VERSION : 0.1
   VAR_INPUT
      "array" : Variant;
   END_VAR
   VAR_TEMP
      status : DInt;
      ret : UDInt;
   END_VAR
BEGIN
   #ret := CountOfElements(#array);
   #"Array.Any.Length" := #ret;
END_FUNCTION

FUNCTION "Get Station Index From Id" : Int   // FC106, SCL
{ S7_Optimized_Access := 'TRUE' }
VERSION : 0.1
   VAR_INPUT
      line_name : WString;
      drop_zone : USInt;
      stns : "Station: All Stations";
   END_VAR
   VAR_TEMP
      i : Int;
      ret : Int;
   END_VAR
BEGIN
   REGION "MATCH LINE NAME AND DROP ZONE"
       FOR #i := 0 TO "STATION_COUNT" DO
           IF #line_name = #stns.stn[#i].id.lineName THEN
               IF #drop_zone = #stns.stn[#i].id.dropZone THEN
                   #ret := #i;
                   EXIT;
               END_IF;
           END_IF;
       END_FOR;
   END_REGION


   REGION "RETURN"
       #"Get Station Index From Id" := #ret;
   END_REGION
END_FUNCTION

FUNCTION "Array.Int.Fill" : Void   // FC109, SCL
{ S7_Optimized_Access := 'TRUE' }
VERSION : 0.1
   VAR_INPUT
      value : Int;
   END_VAR
   VAR_IN_OUT
      int_array : Array[*] of Int;
   END_VAR
   VAR_TEMP
      _i : DInt;
      _length : DInt;
   END_VAR
BEGIN
   REGION "GET LENGHT"
       #_length := UDINT_TO_DINT("Array.Any.Length"(#int_array));
       #_length -= 1;
   END_REGION


   REGION "FILL LENGTH WITH BYTE IN"
       FOR #_i := 0 TO #_length DO
           #int_array[#_i] := #value;
       END_FOR;
   END_REGION
END_FUNCTION

FUNCTION "Array.DInt.Is_Element" : Bool   // FC111, SCL
{ S7_Optimized_Access := 'TRUE' }
VERSION : 0.1
   VAR_INPUT
      dint_array : Array[*] of DInt;
      search_term : DInt;
   END_VAR
   VAR_TEMP
      _i : DInt;
      _length : DInt;
   END_VAR
BEGIN
   REGION "LOCAL VARIABLES"
       #_length := UDINT_TO_DINT("Array.Any.Length"(#dint_array)) - 1;
   END_REGION


   REGION "SEARCH ARRAY"
       FOR #_i := 0 TO #_length DO
           IF #dint_array[#_i] <> #search_term THEN
               CONTINUE;
           END_IF;
           #"Array.DInt.Is_Element" := TRUE;
           RETURN;
       END_FOR;
   END_REGION


   REGION "NOT FOUND"
       #"Array.DInt.Is_Element" := FALSE;
       RETURN;
   END_REGION
END_FUNCTION

FUNCTION "Array.Int.Collapse" : Void   // FC114, SCL
{ S7_Optimized_Access := 'TRUE' }
VERSION : 0.1
   VAR_INPUT
      null_value : Int;   // value that indicates null data
   END_VAR
   VAR_IN_OUT
      int_array : Variant;
   END_VAR
   VAR_TEMP
      i : Int;
      j : Int;
      len_int : Int;
      len_udint : UDInt;
      status : Int;
      t_int_array : Array[0..999] of Int;
   END_VAR
BEGIN
   REGION "COPY TO LOCAL MEMORY"
       #len_udint := CountOfElements(#int_array);
       #len_int := UDINT_TO_INT(#len_udint) - 1;
       #status := MOVE_BLK_VARIANT(SRC := #int_array,
                                   COUNT := #len_udint,
                                   SRC_INDEX := 0,
                                   DEST_INDEX := 0,
                                   DEST => #t_int_array);
   END_REGION

   REGION "COLLAPSE IN PLACE"
       FOR #i := 0 TO #len_int - 1 DO
           IF #t_int_array[#i] = #null_value THEN
               FOR #j := #i + 1 TO #len_int DO
                   IF #t_int_array[#j] <> #null_value THEN
                       #t_int_array[#i] := #t_int_array[#j];
                       #t_int_array[#j] := #null_value;
                       EXIT;
                   END_IF;
               END_FOR;
           END_IF;
       END_FOR;
   END_REGION

   REGION "RETURN"
       #status := MOVE_BLK_VARIANT(SRC := #t_int_array,
                                   COUNT := #len_udint,
                                   SRC_INDEX := 0,
                                   DEST_INDEX := 0,
                                   DEST => #int_array);
   END_REGION
END_FUNCTION

FUNCTION "Array.Int.Count" : Int   // FC115, SCL
{ S7_Optimized_Access := 'TRUE' }
VERSION : 0.1
   VAR_INPUT
      null_value : Int;
      "array" : Variant;
   END_VAR
   VAR_TEMP
      count : Int;
      i : Int;
      len_int : Int;
      len_udint : UDInt;
      status : Int;
      t_array : Array[0..999] of Int;
   END_VAR
BEGIN
   REGION "NOTES"
       (*
       returns the number of valid elements in a collapsed int array
       *)
   END_REGION


   REGION "COPY TO LOCAL"
       #len_udint := CountOfElements(#array);
       #len_int := UDINT_TO_INT(#len_udint) - 1;
       #status := MOVE_BLK_VARIANT(SRC := #array,
                                   COUNT := #len_udint,
                                   SRC_INDEX := 0,
                                   DEST_INDEX := 0,
                                   DEST => #t_array);
   END_REGION


   REGION "SCAN FOR FIRST NULL"
       FOR #i := 0 TO #len_int DO
           IF #t_array[#i] = #null_value THEN
               EXIT;
           END_IF;
           IF #t_array[#i] <> #null_value THEN
               #count += 1;
           END_IF;
       END_FOR;
   END_REGION


   REGION "RETURN"
       #"Array.Int.Count" := #count;
   END_REGION
END_FUNCTION

FUNCTION "Array.Bool.True_Indices" : Void   // FC120, SCL
{ S7_Optimized_Access := 'TRUE' }
VERSION : 0.1
   VAR_INPUT
      array_of_bool : Array[*] of Bool;   // max 1000 elements
      length : Int;   // necessary because dynamically sized arrays of bool get passed as arrays with size of a multiple of 8
   END_VAR
   VAR_IN_OUT
      list_of_indices : Array[*] of Int;   // max 1000 elements
   END_VAR
   VAR_TEMP
      _i : Int;
      _p_return : Int;
      _resized_bool_array : Array[0..#UBOUND] of Bool;
   END_VAR
   VAR CONSTANT
      UBOUND : Int := 999;
   END_VAR
BEGIN
   REGION "FILL RETURN ARRAY"
       "Array.Int.Fill"(value := "NULL_TOKEN",
                        int_array := #list_of_indices);
   END_REGION


   REGION "COPY TO ARRAY OF STATIC SIZE"
       FOR #_i := 0 TO #length DO
           #_resized_bool_array[#_i] := #array_of_bool[#_i];
       END_FOR;
   END_REGION


   REGION "INSERT INDICES INTO RETURN ARRAY"
       FOR #_i := 0 TO #length DO
           IF #_resized_bool_array[#_i] THEN
               #list_of_indices[#_p_return] := #_i;
               #_p_return += 1;
           END_IF;
       END_FOR;
   END_REGION
END_FUNCTION

FUNCTION "Array.Int.Is_Element" : Bool   // FC121, SCL
{ S7_Optimized_Access := 'TRUE' }
VERSION : 0.1
   VAR_INPUT
      int_array : Array[*] of Int;
      search_term : Int;
   END_VAR
   VAR_TEMP
      _i : Int;
      _length : DInt;
   END_VAR
BEGIN
   REGION "LOCAL VARIABLES"
       #_length := UDINT_TO_DINT("Array.Any.Length"(#int_array)) - 1;
   END_REGION


   REGION "SEARCH ARRAY"
       FOR #_i := 0 TO #_length DO
           IF #int_array[#_i] <> #search_term THEN
               CONTINUE;
           END_IF;
           #"Array.Int.Is_Element" := TRUE;
           RETURN;
       END_FOR;
   END_REGION


   REGION "NOT FOUND"
       #"Array.Int.Is_Element" := FALSE;
       RETURN;
   END_REGION
END_FUNCTION

FUNCTION "Array.DInt.Fill" : Void   // FC131, SCL
{ S7_Optimized_Access := 'TRUE' }
VERSION : 0.1
   VAR_INPUT
      int_in : DInt;
   END_VAR
   VAR_OUTPUT
      array_out : Variant;
   END_VAR
   VAR_TEMP
      i : Int;
      internal_array : Array[0..999] of DInt;
      len_array_out : UDInt;
      status : Int;
   END_VAR
BEGIN
   REGION "GET LENGHT"
       #len_array_out := CountOfElements(#array_out);
   END_REGION


   REGION "FILL LENGTH WITH BYTE IN"
       FOR #i := 0 TO UDINT_TO_INT(#len_array_out) - 1 DO
           #internal_array[#i] := #int_in;
       END_FOR;
   END_REGION


   REGION "RETURN"
       #status := MOVE_BLK_VARIANT(SRC := #internal_array,
                                   COUNT := #len_array_out,
                                   SRC_INDEX := 0,
                                   DEST_INDEX := 0,
                                   DEST => #array_out);
   END_REGION
END_FUNCTION

FUNCTION "Array.Int.Search" : Int   // FC140, SCL
{ S7_Optimized_Access := 'TRUE' }
VERSION : 0.1
   VAR_INPUT
      array_of_int : Variant;   // max upper bound 999
      search_term : Int;
   END_VAR
   VAR_TEMP
      i : Int;
      len_as_udint : UDInt;
      len_as_int : Int;
      ret : Int;
      status : Int;
      t_array : Array[0..999] of Int;
   END_VAR
   // Ret_Val : index of search term. returns -1 if not found.
BEGIN
   REGION "LOCAL VARIABLES"
       #len_as_udint := CountOfElements(#array_of_int);
       #len_as_int := UDINT_TO_INT(#len_as_udint) - 1;
       #status := MOVE_BLK_VARIANT(SRC := #array_of_int,
                                   COUNT := #len_as_udint,
                                   SRC_INDEX := 0,
                                   DEST_INDEX := 0,
                                   DEST => #t_array);
       #ret := -1;
   END_REGION


   REGION "SEARCH ARRAY"
       FOR #i := 0 TO #len_as_int DO
           IF #t_array[#i] = #search_term THEN
               #ret := #i;
               EXIT;
           END_IF;
       END_FOR;
   END_REGION


   REGION "RETURN"
       #"Array.Int.Search" := #ret;
   END_REGION
END_FUNCTION

FUNCTION "Array.Int.Intersect" : Void   // FC141, SCL
{ S7_Optimized_Access := 'TRUE' }
VERSION : 0.1
   VAR_INPUT
      "a" : Variant;   // should be array of int, max 999
      "b" : Variant;   // should be array of int, max 999
      null_value : Int;
   END_VAR
   VAR_OUTPUT
      intersect_array : Variant;   // should be array of int, max 999
   END_VAR
   VAR_TEMP
      i : Int;
      j : Int;
      len_a : Struct
         as_udint : UDInt;
         as_int : Int;
      END_STRUCT;
      len_b : Struct
         as_udint : UDInt;
         as_int : Int;
      END_STRUCT;
      len_longer : Struct
         as_udint : UDInt;
         as_int : Int;
      END_STRUCT;
      len_shorter : Struct
         as_udint : UDInt;
         as_int : Int;
      END_STRUCT;
      t_a : Array[0..#u_bound] of Int;
      p_ret : Int;
      ret : Array[0..#u_bound_double] of Int;
      t_b : Array[0..#u_bound] of Int;
      status : Int;
   END_VAR
   VAR CONSTANT
      u_bound : Int := 999;
      u_bound_double : Int := 1999;
   END_VAR
BEGIN
   REGION "GET LENGTHS"
       #len_a.as_udint := CountOfElements(#a);
       #len_a.as_int := UDINT_TO_INT(#len_a.as_udint) - 1;
       #len_b.as_udint := CountOfElements(#b);
       #len_b.as_int := UDINT_TO_INT(#len_b.as_udint) - 1;
   END_REGION

   REGION "MOVE"
       #status := MOVE_BLK_VARIANT(SRC := #a, COUNT := #len_a.as_udint, SRC_INDEX := 0, DEST_INDEX := 0, DEST => #t_a);
       #status := MOVE_BLK_VARIANT(SRC := #b, COUNT := #len_b.as_udint, SRC_INDEX := 0, DEST_INDEX := 0, DEST => #t_b);
   END_REGION

   REGION "FIND INTERSECT"
       FOR #i := 0 TO #len_a.as_int DO
           IF #t_a[#i] = #null_value THEN
               EXIT;
           END_IF;
           FOR #j := 0 TO #len_b.as_int DO
               IF #t_b[#j] = #null_value THEN
                   EXIT;
               END_IF;
               IF #t_a[#i] = #t_b[#j] THEN
                   #ret[#p_ret] := #t_a[#i];
                   #p_ret += 1;
                   EXIT;
               END_IF;
           END_FOR;
       END_FOR;
   END_REGION

   REGION "RETURN"
       #status := MOVE_BLK_VARIANT(SRC := #ret, COUNT := INT_TO_UDINT(#p_ret - 1), SRC_INDEX := 0, DEST_INDEX := 0, DEST => #intersect_array);
   END_REGION
END_FUNCTION

FUNCTION "Array.DInt.First_Occurance" : DInt   // FC143, SCL
{ S7_Optimized_Access := 'TRUE' }
VERSION : 0.1
   VAR_INPUT
      dint_array : Array[*] of DInt;
      search_term : Int;
   END_VAR
   VAR_TEMP
      _i : DInt;
      _length : UDInt;
   END_VAR
BEGIN
   REGION "NOTES"
       (* 
       This function returns the first occurance of the search term.
       This function meant for use with collapsed arrays.
       See "Array.DInt.Collapse" for collapse functionality.
       *)
   END_REGION


   REGION "GET LENGTH OF INPUT ARRAY"
       #_length := "Array.Any.Length"(#dint_array);
   END_REGION


   REGION "FIND FIRST SEARCH TERM, -1 IF NONE"
       (*
       Its worth noting that "Array.DInt.Is_Element" could return the index of the search term
       as an output, saving the processor some work. 
       The rework is justified by increased encapsulation.
       The time complexity for "Array.DInt.First_Occurance" remains O(n).
       *)
       IF NOT "Array.DInt.Is_Element"(dint_array := #dint_array, search_term := #search_term) THEN
           #"Array.DInt.First_Occurance" := -1;
           RETURN;
       END_IF;
       WHILE #dint_array[#_i] <> #search_term AND DINT_TO_UDINT(#_i) < #_length DO
           #_i += 1;
       END_WHILE;
   END_REGION


   REGION _name_
       #"Array.DInt.First_Occurance" := #_i;
   END_REGION
END_FUNCTION

FUNCTION "Array.DInt.Intersect_Exists" : Bool   // FC144, SCL
{ S7_Optimized_Access := 'TRUE' }
VERSION : 0.1
   VAR_INPUT
      "a" : Variant;   // should be array of dint, max 999
      "b" : Variant;   // should be array of dint, max 999
      null_value : DInt;
   END_VAR
   VAR_TEMP
      i : Int;
      j : Int;
      len_a : Struct
         as_udint : UDInt;
         as_int : Int;
      END_STRUCT;
      len_b : Struct
         as_udint : UDInt;
         as_int : Int;
      END_STRUCT;
      t_a : Array[0..#u_bound] of DInt;
      p_ret : Int;
      ret : Bool;
      t_b : Array[0..#u_bound] of DInt;
      status : Int;
   END_VAR
   VAR CONSTANT
      u_bound : Int := 999;
   END_VAR
BEGIN
   REGION "GET LENGHTS"
       #len_a.as_udint := CountOfElements(#a);
       #len_a.as_int := UDINT_TO_INT(#len_a.as_udint) - 1;
       #len_b.as_udint := CountOfElements(#b);
       #len_b.as_int := UDINT_TO_INT(#len_b.as_udint) - 1;
   END_REGION

   REGION "PERFORM MOVES"
       #status := MOVE_BLK_VARIANT(SRC := #a, COUNT := #len_a.as_udint, SRC_INDEX := 0, DEST_INDEX := 0, DEST => #t_a);
       #status := MOVE_BLK_VARIANT(SRC := #b, COUNT := #len_b.as_udint, SRC_INDEX := 0, DEST_INDEX := 0, DEST => #t_b);
   END_REGION


   REGION "SEARCH FOR ANY MATCHING ELEMENT"
       FOR #i := 0 TO #len_a.as_int DO

           REGION "SKIP NULL VALUES"
               IF #t_a[#i] = #null_value THEN
                   CONTINUE;
               END_IF;
           END_REGION

           REGION "INNER LOOP"
               FOR #j := 0 TO #len_b.as_int DO

                   REGION "SKIP NULL VALUES"
                       IF #t_b[#j] = #null_value THEN
                           CONTINUE;
                       END_IF;
                   END_REGION

                   REGION "SET RETURN VALUE ON MATCH"
                       IF #t_a[#i] = #t_b[#j] THEN
                           #ret := TRUE;
                           EXIT;
                       END_IF;
                   END_REGION

               END_FOR;
           END_REGION

           REGION "EXIT OUTTER LOOP IF MATCH FOUND"
               IF #ret THEN
                   EXIT;
               END_IF;
           END_REGION

       END_FOR;
   END_REGION

   REGION "RETURN"
       #"Array.DInt.Intersect_Exists" := #ret;
   END_REGION
END_FUNCTION

FUNCTION "Array.DInt.Intersect" : Void   // FC145, SCL
{ S7_Optimized_Access := 'TRUE' }
VERSION : 0.1
   VAR_INPUT
      "a" : Variant;   // should be array of dint, max 999
      "b" : Variant;   // should be array of dint, max 999
      null_value : DInt;
   END_VAR
   VAR_OUTPUT
      intersect_array : Variant;   // should be array of dint, max 999
   END_VAR
   VAR_TEMP
      i : Int;
      j : Int;
      len_a : Struct
         as_udint : UDInt;
         as_int : Int;
      END_STRUCT;
      len_b : Struct
         as_udint : UDInt;
         as_int : Int;
      END_STRUCT;
      t_a : Array[0..#u_bound] of DInt;
      p_ret : Int;
      ret : Array[0..#u_bound_double] of DInt;
      t_b : Array[0..#u_bound] of DInt;
      status : Int;
   END_VAR
   VAR CONSTANT
      u_bound : Int := 999;
      u_bound_double : Int := 1999;
   END_VAR
BEGIN
   REGION "GET LENGTHS"
       #len_a.as_udint := CountOfElements(#a);
       #len_a.as_int := UDINT_TO_INT(#len_a.as_udint) - 1;
       #len_b.as_udint := CountOfElements(#b);
       #len_b.as_int := UDINT_TO_INT(#len_b.as_udint) - 1;
   END_REGION

   REGION "MOVE"
       #status := MOVE_BLK_VARIANT(SRC := #a, COUNT := #len_a.as_udint, SRC_INDEX := 0, DEST_INDEX := 0, DEST => #t_a);
       #status := MOVE_BLK_VARIANT(SRC := #b, COUNT := #len_b.as_udint, SRC_INDEX := 0, DEST_INDEX := 0, DEST => #t_b);
   END_REGION

   REGION "FIND INTERSECT"
       FOR #i := 0 TO #len_a.as_int DO
           IF #t_a[#i] = #null_value THEN
               EXIT;
           END_IF;
           FOR #j := 0 TO #len_b.as_int DO
               IF #t_b[#j] = #null_value THEN
                   EXIT;
               END_IF;
               IF #t_a[#i] = #t_b[#j] THEN
                   #ret[#p_ret] := #t_a[#i];
                   #p_ret += 1;
                   EXIT;
               END_IF;
           END_FOR;
       END_FOR;
   END_REGION

   REGION "RETURN"
       #status := MOVE_BLK_VARIANT(SRC := #ret, COUNT := INT_TO_UDINT(#p_ret - 1), SRC_INDEX := 0, DEST_INDEX := 0, DEST => #intersect_array);
   END_REGION
END_FUNCTION

FUNCTION "Array.WString.Is_Element" : Bool   // FC207, SCL
{ S7_Optimized_Access := 'TRUE' }
VERSION : 0.1
   VAR_INPUT
      search_term : WString;
      search_array : Array[*] of WString[1];
   END_VAR
   VAR_TEMP
      _i : Int;
      _length_search_array : UDInt;
   END_VAR
BEGIN
   #_length_search_array := "Array.Any.Length"(#search_array);
   FOR #_i := 0 TO UDINT_TO_INT(#_length_search_array - 1) DO
       IF #search_term = #search_array[#_i] THEN
           #"Array.WString.Is_Element" := TRUE;
           RETURN;
       END_IF;
   END_FOR;
   #"Array.WString.Is_Element" := FALSE;
END_FUNCTION

FUNCTION "Array.Int.First_Occurance" : DInt   // FC220, SCL
{ S7_Optimized_Access := 'TRUE' }
VERSION : 0.1
   VAR_INPUT
      int_array : Array[*] of Int;
      search_term : Int;
   END_VAR
   VAR_TEMP
      _i : DInt;
      _length : UDInt;
   END_VAR
BEGIN
   REGION "NOTES"
       (* 
       This function returns the first occurance of the search term.
       This function meant for use with collapsed arrays.
       See "Array.Int.Collapse" for collapse functionality.
       *)
   END_REGION


   REGION "GET LENGTH OF INPUT ARRAY"
       #_length := "Array.Any.Length"(#int_array);
   END_REGION


   REGION "FIND FIRST SEARCH TERM, -1 IF NONE"
       (*
       Its worth noting that "Array.Int.Is_Element" could return the index of the search term
       as an output, saving the processor some work. 
       The rework is justified by increased encapsulation.
       The time complexity for "Array.Int.First_Occurance" remains O(n).
       *)
       IF NOT "Array.Int.Is_Element"(int_array := #int_array, search_term := #search_term) THEN
           #"Array.Int.First_Occurance" := -1;
           RETURN;
       END_IF;
       WHILE #int_array[#_i] <> #search_term AND DINT_TO_UDINT(#_i) < #_length DO
           #_i += 1;
       END_WHILE;
   END_REGION


   REGION _name_
       #"Array.Int.First_Occurance" := #_i;
   END_REGION
END_FUNCTION

FUNCTION "Array.WString.Fill" : Void   // FC243, SCL
{ S7_Optimized_Access := 'TRUE' }
VERSION : 0.1
   VAR_INPUT
      value : WString;
   END_VAR
   VAR_IN_OUT
      "array" : Array[*] of WString;
   END_VAR
   VAR_TEMP
      _length : Int;
      _i : Int;
   END_VAR
BEGIN
   #_length := UDINT_TO_INT("Array.Any.Length"(#array)) - 1;
   FOR #_i := 0 TO #_length DO
       #array[#_i] := #value;
   END_FOR;
   RETURN;
END_FUNCTION

FUNCTION "Array.WString.Search" : Int   // FC244, SCL
{ S7_Optimized_Access := 'TRUE' }
VERSION : 0.1
   VAR_INPUT
      "array" : Array[*] of WString;
      search_term : WString;
   END_VAR
   VAR_TEMP
      _i : Int;
      _length : Int;
   END_VAR
   // Ret_Val : index of search term. returns -1 if not found.
BEGIN
   REGION "SEARCH ARRAY"    
       #_length := UDINT_TO_INT("Array.Any.Length"(#array)) - 1;
       FOR #_i := 0 TO #_length DO
           IF #array[#_i] = #search_term THEN
               #"Array.WString.Search" := #_i;
               RETURN;
           END_IF;
       END_FOR;
   END_REGION

   REGION "RETURN"
       #"Array.WString.Search" := "NULL_TOKEN";
       RETURN;
   END_REGION
END_FUNCTION

FUNCTION "Array.Char.Search" : Int   // FC266, SCL
{ S7_Optimized_Access := 'TRUE' }
VERSION : 0.1
   VAR_INPUT
      "array" : Array[*] of Char;   // max upper bound 999
      search_term : Char;
   END_VAR
   VAR_TEMP
      _i : Int;
      _length : Int;
   END_VAR
   // Ret_Val : index of search term. returns -1 if not found.
BEGIN
   REGION "GET LENGTH"
       #_length := UDINT_TO_INT("Array.Any.Length"(#array)) - 1;
   END_REGION


   REGION "SEARCH ARRAY"
       FOR #_i := 0 TO #_length DO
           IF #array[#_i] = #search_term THEN
               #"Array.Char.Search" := #_i;
               EXIT;
           END_IF;
       END_FOR;
   END_REGION


   REGION "RETURN"
       #"Array.Char.Search" := "NULL_TOKEN";
   END_REGION
END_FUNCTION

FUNCTION "Array.WString.Reverse" : Void   // FC270, SCL
{ S7_Optimized_Access := 'TRUE' }
VERSION : 0.1
   VAR_INPUT
      null_token : WString;
   END_VAR
   VAR_IN_OUT
      wstring_array : Array[*] of WString;
   END_VAR
   VAR_TEMP
      _has_data_count : Int;
      _i : Int;
      _p_swap : Int;
      _temp : WString;
   END_VAR
   VAR CONSTANT
      NOT_FOUND : Int := -1;
   END_VAR
BEGIN
   REGION "CHECK FOR FIRST EMPTY POSITION"
       #_has_data_count := "Array.WString.Search"(array := #wstring_array,
                                                  search_term := #null_token);
   END_REGION


   REGION "EXIT ON EMPTY ARRAY"
       IF #_has_data_count = 0 THEN
           RETURN;
       END_IF;
   END_REGION


   REGION "ARRAY IS FULL"
       IF #_has_data_count = #NOT_FOUND THEN
           #_has_data_count := UDINT_TO_INT("Array.Any.Length"(#wstring_array));
       END_IF;
   END_REGION


   REGION "ADJUST TO ZERO INDEX"
       #_has_data_count -= 1;
   END_REGION


   REGION "SWAP ELEMENTS"
       FOR #_i := 0 TO #_has_data_count / 2 DO
           #_p_swap := #_has_data_count - #_i;
           #_temp := #wstring_array[#_i];
           #wstring_array[#_i] := #wstring_array[#_p_swap];
           #wstring_array[#_p_swap] := #_temp;
       END_FOR;
   END_REGION


   REGION "DONE"
       RETURN;
   END_REGION
END_FUNCTION

// folder: Utilities/Bool

FUNCTION "Bool.Animate" : USInt   // FC9, SCL
{ S7_Optimized_Access := 'TRUE' }
VERSION : 0.1
   VAR_INPUT
      true_color : USInt;
      false_color : USInt;
      evaluation_signal : Bool;
   END_VAR
   VAR_TEMP
      animate : USInt;
   END_VAR
BEGIN
   REGION "FALSE COLOR"
       IF NOT #evaluation_signal THEN
           #animate := #false_color;
       END_IF;
   END_REGION

   REGION "TRUE COLOR"
       IF #evaluation_signal THEN
           #animate := #true_color;
       END_IF;
   END_REGION

   REGION "FUNCTION RETURN"
       #"Bool.Animate" := #animate;
   END_REGION
END_FUNCTION

FUNCTION "Bool.Rising_Edge" : Bool   // FC177, SCL
{ S7_Optimized_Access := 'TRUE' }
VERSION : 0.1
   VAR_INPUT
      signal : Bool;
      old_signal : Bool;
   END_VAR
BEGIN
   #"Bool.Rising_Edge" := #signal AND NOT #old_signal;
END_FUNCTION

FUNCTION "Bool.Falling_Edge" : Bool   // FC178, SCL
{ S7_Optimized_Access := 'TRUE' }
VERSION : 0.1
   VAR_INPUT
      signal : Bool;
      old_signal : Bool;
   END_VAR
BEGIN
   #"Bool.Falling_Edge" := NOT #signal AND #old_signal;
END_FUNCTION

// folder: Utilities/DInt

FUNCTION "Pointer Calc: KP8 Labels" : Int   // FC25, SCL
{ S7_Optimized_Access := 'TRUE' }
VERSION : 0.1
   VAR_INPUT
      index : Int;
   END_VAR
   VAR_TEMP
      val : Int;
   END_VAR
BEGIN
   IF #index >= 4 THEN
       #val := 7 - (#index - 4) * 2;
   END_IF;

   IF #index <= 3 THEN
       #val := 8 - #index * 2;
   END_IF;

   #"Pointer Calc: KP8 Labels" := #val;
END_FUNCTION

FUNCTION "DInt.Clip.Maximum" : DInt   // FC224, SCL
{ S7_Optimized_Access := 'TRUE' }
VERSION : 0.1
   VAR_INPUT
      value : DInt;
      maximum : DInt;
   END_VAR
BEGIN
   IF #value > #maximum THEN
       #"DInt.Clip.Maximum" := #maximum;
       RETURN;
   END_IF;
   #"DInt.Clip.Maximum" := #value;
END_FUNCTION

FUNCTION "DInt.Clip.Minimum" : DInt   // FC225, SCL
{ S7_Optimized_Access := 'TRUE' }
VERSION : 0.1
   VAR_INPUT
      value : DInt;
      minimum : DInt;
   END_VAR
BEGIN
   IF #value < #minimum THEN
       #"DInt.Clip.Minimum" := #minimum;
       RETURN;
   END_IF;
   #"DInt.Clip.Minimum" := #value;
END_FUNCTION

FUNCTION "DInt.Clip.Range" : DInt   // FC227, SCL
{ S7_Optimized_Access := 'TRUE' }
VERSION : 0.1
   VAR_INPUT
      value : DInt;
      maximum : DInt;
      minimum : DInt;
   END_VAR
   VAR_TEMP
      _return : DInt;
   END_VAR
BEGIN
   #_return := #value;
   #_return := "DInt.Clip.Maximum"(value := #value, maximum := #minimum);
   #_return := "DInt.Clip.Minimum"(value := #value, minimum := #minimum);
   #"DInt.Clip.Range" := #_return;
END_FUNCTION

// folder: Utilities/Int

FUNCTION "Int.Value_Change" : Bool   // FC179, SCL
{ S7_Optimized_Access := 'TRUE' }
VERSION : 0.1
   VAR_INPUT
      value : Int;
      old_value : Int;
   END_VAR
BEGIN
   #"Int.Value_Change" := #value <> #old_value;
END_FUNCTION

FUNCTION "Int.Clip.Minimum" : Int   // FC222, SCL
{ S7_Optimized_Access := 'TRUE' }
VERSION : 0.1
   VAR_INPUT
      value : Int;
      minimum : Int;
   END_VAR
BEGIN
   IF #value < #minimum THEN
       #"Int.Clip.Minimum" := #minimum;
       RETURN;
   END_IF;
   #"Int.Clip.Minimum" := #value;
END_FUNCTION

FUNCTION "Int.Clip.Maximum" : Int   // FC223, SCL
{ S7_Optimized_Access := 'TRUE' }
VERSION : 0.1
   VAR_INPUT
      value : Int;
      maximum : Int;
   END_VAR
BEGIN
   IF #value > #maximum THEN
       #"Int.Clip.Maximum" := #maximum;
       RETURN;
   END_IF;
   #"Int.Clip.Maximum" := #value;
END_FUNCTION

FUNCTION "Int.Clip.Range" : Int   // FC226, SCL
{ S7_Optimized_Access := 'TRUE' }
VERSION : 0.1
   VAR_INPUT
      value : Int;
      maximum : Int;
      minimum : Int;
   END_VAR
   VAR_TEMP
      _return : Int;
   END_VAR
BEGIN
   #_return := #value;
   #_return := "Int.Clip.Maximum"(value := #_return, maximum := #maximum);
   #_return := "Int.Clip.Minimum"(value:=#_return, minimum:=#minimum);
   #"Int.Clip.Range" := #_return;
END_FUNCTION

// folder: Utilities/NavBar

FUNCTION_BLOCK "NavBar: Top"   // FB31, SCL
{ S7_Optimized_Access := 'TRUE' }
VERSION : 0.1
   VAR_INPUT
      hide : Bool;
      TABLE_LENGTH : DInt;
   END_VAR
   VAR_IN_OUT
      interface : "Push Button Data";
      first_row : DInt;
   END_VAR
   VAR
      "Get Button Feedback" : "Push Button: State Changes";
   END_VAR
   VAR_TEMP
      feedback : "Push Button Data: State Change Data";
   END_VAR
BEGIN
   REGION "PROCESS USER INPUT"
       #"Get Button Feedback"(interface := #interface,
                              state_changes := #feedback);
   END_REGION

   REGION "ANIMATIONS"

       REGION "COLOR"
           #interface.animate := "Bool.Animate"(true_color := "GREEN_LIGHT_BACKGROUND",
                                                false_color := "GRAY_BACKGROUND",
                                                evaluation_signal := #feedback.actuate.actual);
       END_REGION

       REGION "VISIBILITY"
           #interface.visible := NOT #hide;
       END_REGION

       REGION "ENABLED STATE"
           #interface.enable := NOT #hide;
       END_REGION

   END_REGION

   REGION "SET FIRST ROW"
       IF #feedback.actuate.rising THEN
           #first_row := 0;
       END_IF;
   END_REGION
END_FUNCTION_BLOCK

FUNCTION_BLOCK "NavBar: Bottom"   // FB32, SCL
{ S7_Optimized_Access := 'TRUE' }
VERSION : 0.1
   VAR_INPUT
      hide : Bool;
      TABLE_LENGTH : DInt;
      VISIBLE_ROW_COUNT : DInt;
   END_VAR
   VAR_IN_OUT
      interface : "Push Button Data";
      first_row : DInt;
   END_VAR
   VAR
      "Get Button Feedback" : "Push Button: State Changes";
   END_VAR
   VAR_TEMP
      feedback : "Push Button Data: State Change Data";
   END_VAR
BEGIN
   REGION "PROCESS USER INPUT"
       #"Get Button Feedback"(interface := #interface,
                              state_changes := #feedback);
   END_REGION

   REGION "ANIMATIONS"

       REGION "COLOR"
           #interface.animate := "Bool.Animate"(true_color := "GREEN_LIGHT_BACKGROUND",
                                                false_color := "GRAY_BACKGROUND",
                                                evaluation_signal := #feedback.actuate.actual);
       END_REGION

       REGION "VISIBILITY"
           #interface.visible := NOT #hide;
       END_REGION

       REGION "ENABLED STATE"
           #interface.enable := NOT #hide;
       END_REGION

   END_REGION


   REGION "SET FIRST ROW"
       IF #feedback.actuate.rising THEN
           #first_row := #TABLE_LENGTH - #VISIBLE_ROW_COUNT;
       END_IF;
   END_REGION
END_FUNCTION_BLOCK

FUNCTION_BLOCK "NavBar: Page Up"   // FB36, SCL
{ S7_Optimized_Access := 'TRUE' }
VERSION : 0.1
   VAR_INPUT
      hide : Bool;
      TABLE_LENGTH : DInt;
      VISIBLE_ROW_COUNT : DInt;
   END_VAR
   VAR_IN_OUT
      interface : "Push Button Data";
      first_row : DInt;
   END_VAR
   VAR
      "Get Button Feedback" : "Push Button: State Changes";
   END_VAR
   VAR_TEMP
      feedback : "Push Button Data: State Change Data";
   END_VAR
BEGIN
   REGION "PROCESS USER INPUT"
       #"Get Button Feedback"(interface := #interface,
                              state_changes := #feedback);
   END_REGION

   REGION "ANIMATIONS"

       REGION "COLOR"
           #interface.animate := "Bool.Animate"(true_color := "GREEN_LIGHT_BACKGROUND",
                                                false_color := "GRAY_BACKGROUND",
                                                evaluation_signal := #feedback.actuate.actual);
       END_REGION

       REGION "VISIBILITY"
           #interface.visible := NOT #hide;
       END_REGION

       REGION "ENABLED STATE"
           #interface.enable := NOT #hide;
       END_REGION

   END_REGION

   REGION "SET FIRST ROW"
       IF #feedback.actuate.rising THEN
           #first_row := "NavBar: Private: First Row"(first_row := #first_row,
                                                      offset := -1 * (#VISIBLE_ROW_COUNT + 1),
                                                      TABLE_LENGTH := #TABLE_LENGTH);
       END_IF;
   END_REGION
END_FUNCTION_BLOCK

FUNCTION_BLOCK "NavBar: Page Down"   // FB37, SCL
{ S7_Optimized_Access := 'TRUE' }
VERSION : 0.1
   VAR_INPUT
      hide : Bool;
      TABLE_LENGTH : DInt;
      VISIBLE_ROW_COUNT : DInt;
   END_VAR
   VAR_IN_OUT
      interface : "Push Button Data";
      first_row : DInt;
   END_VAR
   VAR
      "Get Button Feedback" : "Push Button: State Changes";
   END_VAR
   VAR_TEMP
      feedback : "Push Button Data: State Change Data";
   END_VAR
BEGIN
   REGION "PROCESS USER INPUT"
       #"Get Button Feedback"(interface := #interface,
                              state_changes := #feedback);
   END_REGION

   REGION "ANIMATIONS"

       REGION "COLOR"
           #interface.animate := "Bool.Animate"(true_color := "GREEN_LIGHT_BACKGROUND",
                                                false_color := "GRAY_BACKGROUND",
                                                evaluation_signal := #feedback.actuate.actual);
       END_REGION

       REGION "VISIBILITY"
           #interface.visible := NOT #hide;
       END_REGION

       REGION "ENABLED STATE"
           #interface.enable := NOT #hide;
       END_REGION

   END_REGION

   REGION "SET FIRST ROW"
       IF #feedback.actuate.rising THEN
           #first_row := "NavBar: Private: First Row"(first_row := #first_row,
                                                      offset := #VISIBLE_ROW_COUNT + 1,
                                                      TABLE_LENGTH := #TABLE_LENGTH);
       END_IF;
   END_REGION
END_FUNCTION_BLOCK

FUNCTION_BLOCK "NavBar: Line Down"   // FB38, SCL
{ S7_Optimized_Access := 'TRUE' }
VERSION : 0.1
   VAR_INPUT
      hide : Bool;
      TABLE_LENGTH : DInt;
   END_VAR
   VAR_IN_OUT
      interface : "Push Button Data";
      first_row : DInt;
   END_VAR
   VAR
      "Get Button Feedback" : "Push Button: State Changes";
   END_VAR
   VAR_TEMP
      feedback : "Push Button Data: State Change Data";
   END_VAR
BEGIN
   REGION "PROCESS USER INPUT"
       #"Get Button Feedback"(interface := #interface,
                              state_changes := #feedback);
   END_REGION

   REGION "ANIMATIONS"

       REGION "COLOR"
           #interface.animate := "Bool.Animate"(true_color := "GREEN_LIGHT_BACKGROUND",
                                                false_color := "GRAY_BACKGROUND",
                                                evaluation_signal := #feedback.actuate.actual);
       END_REGION

       REGION "VISIBILITY"
           #interface.visible := NOT #hide;
       END_REGION

       REGION "ENABLED STATE"
           #interface.enable := NOT #hide;
       END_REGION

   END_REGION

   REGION "SET FIRST ROW"
       IF #feedback.actuate.rising THEN
           #first_row := "NavBar: Private: First Row"(first_row := #first_row,
                                                      offset := 1,
                                                      TABLE_LENGTH := #TABLE_LENGTH);
       END_IF;
   END_REGION
END_FUNCTION_BLOCK

FUNCTION_BLOCK "NavBar: Line Up"   // FB39, SCL
{ S7_Optimized_Access := 'TRUE' }
VERSION : 0.1
   VAR_INPUT
      hide : Bool;
      TABLE_LENGTH : DInt;
   END_VAR
   VAR_IN_OUT
      interface : "Push Button Data";
      first_row : DInt;
   END_VAR
   VAR
      "Get Button Feedback" : "Push Button: State Changes";
   END_VAR
   VAR_TEMP
      feedback : "Push Button Data: State Change Data";
   END_VAR
BEGIN
   REGION "PROCESS USER INPUT"
       #"Get Button Feedback"(interface := #interface,
                              state_changes := #feedback);
   END_REGION

   REGION "ANIMATIONS"

       REGION "COLOR"
           #interface.animate := "Bool.Animate"(true_color := "GREEN_LIGHT_BACKGROUND",
                                                false_color := "GRAY_BACKGROUND",
                                                evaluation_signal := #feedback.actuate.actual);
       END_REGION

       REGION "VISIBILITY"
           #interface.visible := NOT #hide;
       END_REGION

       REGION "ENABLED STATE"
           #interface.enable := NOT #hide;
       END_REGION

   END_REGION

   REGION "SET FIRST ROW"
       IF #feedback.actuate.rising THEN
           #first_row := "NavBar: Private: First Row"(first_row := #first_row,
                                                      offset := -1,
                                                      TABLE_LENGTH := #TABLE_LENGTH);
       END_IF;
   END_REGION
END_FUNCTION_BLOCK

FUNCTION_BLOCK "NavBar"   // FB40, SCL
{ S7_Optimized_Access := 'TRUE' }
VERSION : 0.1
   VAR_INPUT
      hide : Bool;
      TABLE_LENGTH : DInt := 49;
      VISIBLE_ROW_COUNT : DInt := 2;
   END_VAR
   VAR_IN_OUT
      interface : "Nav Bar Data";
      first_row : DInt;
   END_VAR
   VAR
      Top : "NavBar: Top";
      "Page Up" : "NavBar: Page Up";
      "Line Up" : "NavBar: Line Up";
      "Line Down" : "NavBar: Line Down";
      "Page Down" : "NavBar: Page Down";
      Bottom : "NavBar: Bottom";
   END_VAR
BEGIN
   REGION "BUFFER IN"
       "NavBar: Map HMI to PLC"(hmi := #interface.hmi,
                                plc := #interface.plc);
   END_REGION

   REGION "NAVBAR TOP "
       #Top(hide := #hide,
            TABLE_LENGTH := #TABLE_LENGTH,
            interface := #interface.plc.top,
            first_row := #first_row);
   END_REGION

   REGION "PAGE UP"
       #"Page Up"(hide := #hide,
                  TABLE_LENGTH := #TABLE_LENGTH,
                  VISIBLE_ROW_COUNT := #VISIBLE_ROW_COUNT,
                  interface := #interface.plc.pageUp,
                  first_row := #first_row);
   END_REGION

   REGION "LINE UP"
       #"Line Up"(hide := #hide,
                  TABLE_LENGTH := #TABLE_LENGTH,
                  interface := #interface.plc.lineUp,
                  first_row := #first_row);
   END_REGION

   REGION "LINE DOWN"
       #"Line Down"(hide := #hide,
                    TABLE_LENGTH := #TABLE_LENGTH,
                    interface := #interface.plc.lineDown,
                    first_row := #first_row);
   END_REGION

   REGION "PAGE DOWN"
       #"Page Down"(hide := #hide,
                    TABLE_LENGTH := #TABLE_LENGTH,
                    VISIBLE_ROW_COUNT := #VISIBLE_ROW_COUNT,
                    interface := #interface.plc.pageDown,
                    first_row := #first_row);
   END_REGION

   REGION "BOTTOM"
       #Bottom(hide := #hide,
               TABLE_LENGTH := #TABLE_LENGTH,
               VISIBLE_ROW_COUNT := #VISIBLE_ROW_COUNT,
               interface := #interface.plc.bottom,
               first_row := #first_row);
   END_REGION

   REGION "BUFFER OUT"
       "NavBar: Map PLC to HMI"(plc := #interface.plc,
                                hmi := #interface.hmi);
   END_REGION
END_FUNCTION_BLOCK

FUNCTION "NavBar: Map HMI to PLC" : Void   // FC98, SCL
{ S7_Optimized_Access := 'TRUE' }
VERSION : 0.1
   VAR_INPUT
      hmi : "Nav Bar Data: HMI";
   END_VAR
   VAR_IN_OUT
      plc : "Nav Bar Data: PLC";
   END_VAR
BEGIN
   REGION "NOTES"
       // mapping is necessary because hmi faceplate data structures
       // cannot consist of embedded udts
   END_REGION


   REGION "TOP"
       #plc.top.actuate := #hmi.top_actuate;
       #plc.top.animate := #hmi.top_animate;
       #plc.top.enable := #hmi.top_enable;
       #plc.top.label := #hmi.top_label;
       #plc.top.listSelect := #hmi.top_list_select;
       #plc.top.visible := #hmi.top_visible;
   END_REGION


   REGION "PAGE UP"
       #plc.pageUp.actuate := #hmi.page_up_actuate;
       #plc.pageUp.animate := #hmi.page_up_animate;
       #plc.pageUp.enable := #hmi.page_up_enable;
       #plc.pageUp.label := #hmi.page_up_label;
       #plc.pageUp.listSelect := #hmi.page_up_list_select;
       #plc.pageUp.visible := #hmi.page_up_visible;
   END_REGION


   REGION "LINE UP"
       #plc.lineUp.actuate := #hmi.line_up_actuate;
       #plc.lineUp.animate := #hmi.line_up_animate;
       #plc.lineUp.enable := #hmi.line_up_enable;
       #plc.lineUp.label := #hmi.line_up_label;
       #plc.lineUp.listSelect := #hmi.line_up_list_select;
       #plc.lineUp.visible := #hmi.line_up_visible;
   END_REGION


   REGION "LINE DOWN"
       #plc.lineDown.actuate := #hmi.line_down_actuate;
       #plc.lineDown.animate := #hmi.line_down_animate;
       #plc.lineDown.enable := #hmi.line_down_enable;
       #plc.lineDown.label := #hmi.line_down_label;
       #plc.lineDown.listSelect := #hmi.line_down_list_select;
       #plc.lineDown.visible := #hmi.line_down_visible;
   END_REGION


   REGION "PAGE DOWN"
       #plc.pageDown.actuate := #hmi.page_down_actuate;
       #plc.pageDown.animate := #hmi.page_down_animate;
       #plc.pageDown.enable := #hmi.page_down_enable;
       #plc.pageDown.label := #hmi.page_down_label;
       #plc.pageDown.listSelect := #hmi.page_down_list_select;
       #plc.pageDown.visible := #hmi.page_down_visible;
   END_REGION


   REGION "BOTTOM"
       #plc.bottom.actuate := #hmi.bottom_actuate;
       #plc.bottom.animate := #hmi.bottom_animate;
       #plc.bottom.enable := #hmi.bottom_enable;
       #plc.bottom.label := #hmi.bottom_label;
       #plc.bottom.listSelect := #hmi.bottom_list_select;
       #plc.bottom.visible := #hmi.bottom_visible;
   END_REGION
END_FUNCTION

FUNCTION "NavBar: Map PLC to HMI" : Void   // FC99, SCL
{ S7_Optimized_Access := 'TRUE' }
VERSION : 0.1
   VAR_INPUT
      plc : "Nav Bar Data: PLC";
   END_VAR
   VAR_IN_OUT
      hmi : "Nav Bar Data: HMI";
   END_VAR
BEGIN
   REGION "NOTES"
       // mapping is necessary because hmi faceplate data structures
       // cannot consist of embedded udts
   END_REGION


   REGION "TOP"
       //#hmi.top_actuate := #plc.top.actuate;
       #hmi.top_animate := #plc.top.animate;
       #hmi.top_enable := #plc.top.enable;
       #hmi.top_label := #plc.top.label;
       #hmi.top_list_select := #plc.top.listSelect;
       #hmi.top_visible := #plc.top.visible;
   END_REGION


   REGION "PAGE UP"
       //#hmi.page_up_actuate := #plc.pageUp.actuate;
       #hmi.page_up_animate := #plc.pageUp.animate;
       #hmi.page_up_enable := #plc.pageUp.enable;
       #hmi.page_up_label := #plc.pageUp.label;
       #hmi.page_up_list_select := #plc.pageUp.listSelect;
       #hmi.page_up_visible := #plc.pageUp.visible;
   END_REGION


   REGION "LINE UP"
       //#hmi.line_up_actuate := #plc.lineUp.actuate;
       #hmi.line_up_animate := #plc.lineUp.animate;
       #hmi.line_up_enable := #plc.lineUp.enable;
       #hmi.line_up_label := #plc.lineUp.label;
       #hmi.line_up_list_select := #plc.lineUp.listSelect;
       #hmi.line_up_visible := #plc.lineUp.visible;
   END_REGION


   REGION "LINE DOWN"
       //#hmi.line_down_actuate := #plc.lineDown.actuate;
       #hmi.line_down_animate := #plc.lineDown.animate;
       #hmi.line_down_enable := #plc.lineDown.enable;
       #hmi.line_down_label := #plc.lineDown.label;
       #hmi.line_down_list_select := #plc.lineDown.listSelect;
       #hmi.line_down_visible := #plc.lineDown.visible;
   END_REGION


   REGION "PAGE DOWN"
       //#hmi.page_down_actuate := #plc.pageDown.actuate;
       #hmi.page_down_animate := #plc.pageDown.animate;
       #hmi.page_down_enable := #plc.pageDown.enable;
       #hmi.page_down_label := #plc.pageDown.label;
       #hmi.page_down_list_select := #plc.pageDown.listSelect;
       #hmi.page_down_visible := #plc.pageDown.visible;
   END_REGION

   REGION "BOTTOM"
       //#hmi.bottom_actuate := #plc.bottom.actuate;
       #hmi.bottom_animate := #plc.bottom.animate;
       #hmi.bottom_enable := #plc.bottom.enable;
       #hmi.bottom_label := #plc.bottom.label;
       #hmi.bottom_list_select := #plc.bottom.listSelect;
       #hmi.bottom_visible := #plc.bottom.visible;
   END_REGION
END_FUNCTION

FUNCTION "NavBar: Private: First Row" : DInt   // FC180, SCL
{ S7_Optimized_Access := 'TRUE' }
VERSION : 0.1
   VAR_INPUT
      first_row : DInt;
      offset : DInt;
      TABLE_LENGTH : DInt;
   END_VAR
   VAR_TEMP
      ret : DInt;
   END_VAR
BEGIN
   REGION "DESCRIPTION"
       (*
       The new first row of the table is calculated from the offset. 
       Rollover and rollunder are resolved for the first row.
       *)
   END_REGION

   REGION "COPY TO INTERNAL"
       #ret := #first_row + #offset;
   END_REGION

   REGION "ROLLUNDER"
       IF #ret < 0 THEN
           #ret := #ret + #TABLE_LENGTH + 1;
       END_IF;
   END_REGION

   REGION "ROLLOVER"
       IF #ret > #TABLE_LENGTH THEN
           #ret := #ret - #TABLE_LENGTH - 1;
       END_IF;
   END_REGION

   REGION "OUTPUT"
       #"NavBar: Private: First Row" := #ret;
   END_REGION
END_FUNCTION

// folder: Utilities/Part Number

FUNCTION_BLOCK "IO Field: State Changes"   // FB48, SCL
{ S7_Optimized_Access := 'TRUE' }
VERSION : 0.1
   VAR_IN_OUT
      interface : "IO Field Data: Label with Data";
      feedback : "IO Field: State Change Data";
   END_VAR
   VAR
      old : "IO Field Data: Label with Data";
   END_VAR
BEGIN
   REGION "ANIMATE"
       #feedback.animate.rising := "USInt.Value_Change"(value := #interface.animate,
                                                         old_value := #old.animate);
       #feedback.animate.actual := #interface.animate;
       #feedback.animate.falling := FALSE;     // animate never set to null token 
   END_REGION

   REGION "ENABLE"
       #feedback.enable.rising := "Bool.Rising_Edge"(signal := #interface.enable,
                                                      old_signal := #old.enable);
       #feedback.enable.actual := #interface.enable;
       #feedback.enable.falling := "Bool.Falling_Edge"(signal := #interface.enable,
                                                        old_signal := #old.enable);
   END_REGION

   REGION "INPUT FINISHED"
       #feedback.input_finished.rising := "Bool.Rising_Edge"(signal := #interface.input_finished,
                                                              old_signal := #old.input_finished);
       #feedback.input_finished.actual := #interface.input_finished;
       #feedback.input_finished.falling := "Bool.Falling_Edge"(signal := #interface.input_finished,
                                                                old_signal := #old.input_finished);
   END_REGION

   REGION "VALUE CHANGED"
       #feedback.value.rising := "WString.Rising_Edge"(value := #interface.value,
                                                        old_value := #old.value);
       #feedback.value.actual := #interface.value;
       #feedback.value.falling := "WString.Falling_Edge"(value := #interface.value,
                                                          old_value := #old.value);
   END_REGION

   REGION "VISIBLE"
       #feedback.visible.rising := "Bool.Rising_Edge"(signal := #interface.visible,
                                                       old_signal := #old.visible);
       #feedback.visible.actual := #interface.visible;
       #feedback.visible.falling := "Bool.Falling_Edge"(signal := #interface.visible,
                                                         old_signal := #old.visible);
   END_REGION

   REGION "SAVE OLD VALUES"
       #old := #interface;
   END_REGION
END_FUNCTION_BLOCK

FUNCTION "Part_Number.Parse_Code" : Void   // FC34, SCL
{ S7_Optimized_Access := 'TRUE' }
VERSION : 0.1
   VAR_INPUT
      code : DInt;
   END_VAR
   VAR_OUTPUT
      code_left : DInt;
      code_right : DInt;
   END_VAR
BEGIN
   IF #code > 0 THEN
       #code_left := #code / 1000;
       #code_right := #code - #code / 1000 * 1000;
   ELSE
       #code_left := 0;
       #code_right := 0;
   END_IF;
END_FUNCTION

FUNCTION "Part_Number.Code_to_WString" : WString   // FC37, SCL
{ S7_Optimized_Access := 'TRUE' }
VERSION : 0.1
   VAR_INPUT
      pnLib : "Recipe: PN Text Library";
      pnCode : DInt;
   END_VAR
   VAR_TEMP
      pnLeft : DInt;
      pnRight : DInt;
      output : WString;
   END_VAR
   VAR CONSTANT
      newLine : WString := WSTRING#'$L';
   END_VAR
BEGIN
   REGION "PARSE CODE"
       "Part_Number.Parse_Code"(code := #pnCode,
                                 code_left => #pnLeft,
                                 code_right => #pnRight);
   END_REGION

   REGION "SINGLE LINE PN"
       IF "Part_Number.Is_Single"(#pnCode) THEN
           #output := #pnLib.pnText[#pnLeft];
       END_IF;
   END_REGION

   REGION "DOUBLE LINE PN"
       IF "Part_Number.Is_Double"(#pnCode) THEN
           #output := CONCAT_WSTRING(IN1 := #pnLib.pnText[#pnLeft],
                                     IN2 := #newLine,
                                     IN3 := #pnLib.pnText[#pnRight]);
       END_IF;
   END_REGION

   REGION "OUTPUT"
       #"Part_Number.Code_to_WString" := #output;
   END_REGION
END_FUNCTION

FUNCTION "Part_Number.Is_Double" : Bool   // FC153, SCL
{ S7_Optimized_Access := 'TRUE' }
VERSION : 0.1
   VAR_INPUT
      code : DInt;
   END_VAR
   VAR_TEMP
      code_left : DInt;
      code_right : DInt;
      ret : Bool;
   END_VAR
BEGIN
   REGION "NOTES"
       (*
       Double codes have a non-zero right hand component.
       Structure: XXXYYY
       XXX: left code, used for single and double codes
       YYY: right code, only used for double codes
       Last Edit: 2021-10-07
       *)
   END_REGION

   REGION "PROCESS CODE"
       "Part_Number.Parse_Code"(code := #code,
                                code_left => #code_left,
                                code_right => #code_right);
   END_REGION

   REGION "CHECK FOR DOUBLE CODE"
       IF #code_right > 0 THEN
           #ret := TRUE;
       END_IF;
   END_REGION

   REGION "RETURN" 
       #"Part_Number.Is_Double" := #ret;
   END_REGION
END_FUNCTION

FUNCTION "Part_Number.Is_Single" : Bool   // FC154, SCL
{ S7_Optimized_Access := 'TRUE' }
VERSION : 0.1
   VAR_INPUT
      code : DInt;
   END_VAR
   VAR_TEMP
      code_left : DInt;
      code_right : DInt;
      ret : Bool;
   END_VAR
BEGIN
   REGION "NOTES"
       (*
       Double codes have a non-zero right hand component.
       Structure:
       XXXYYY
       XXX: left code, used for single and double codes
       YYY: right code, only used for double codes
       Last Edit: 2021-10-07
       *)
   END_REGION

   REGION "PROCESS CODE"
       "Part_Number.Parse_Code"(code := #code,
                                code_left => #code_left,
                                code_right => #code_right);
   END_REGION

   REGION "CHECK FOR DOUBLE CODE"
       IF #code_right = 0 THEN
           #ret := TRUE;
       END_IF;
   END_REGION

   REGION "RETURN" 
       #"Part_Number.Is_Single" := #ret;
   END_REGION
END_FUNCTION

FUNCTION "Part_Number.WString_to_Code" : DInt   // FC240, SCL
{ S7_Optimized_Access := 'TRUE' }
VERSION : 0.1
   VAR_INPUT
      part_number : WString;
   END_VAR
   VAR_IN_OUT
      pn_library : "Recipe: PN Text Library";
   END_VAR
   VAR_TEMP
      _in_library : Bool;
      _library_full : Bool;
      _part_numbers : Array[0..1] of WString;
      _partial_pn_code : DInt;
      _pn_count : Int;
      _pn_code : DInt;
   END_VAR
   VAR CONSTANT
      OUT_OF_MEMORY : DInt := 999;
   END_VAR
BEGIN
   REGION "DATA PREP""
       "Part_Number.Split_PNs"(part_number := #part_number,
                               part_numbers := #_part_numbers);
       #_pn_count := "Part_Number.Count_PNs"(#_part_numbers);
   END_REGION


   REGION "NO PART NUMBERS ENTERED"
       IF #_pn_count = 0 THEN
           #"Part_Number.WString_to_Code" := 0;
           RETURN;
       END_IF;
   END_REGION


   REGION "CHECK FIRST PN CODE"
       #_pn_code := "Part_Number_Library.Search"(pn_library := #pn_library,
                                                 search_term := #_part_numbers[0]);
       #_in_library := "Part_Number.In_Library"(#_pn_code);
       #_library_full := "Part_Number_Library.Is_Full"(#pn_library);
   END_REGION


